
screen "MTA-AyudaVentiladores" 1280x800, template "Plantilla"
   GraphicIOField "Campo ES gráfico_6" at 328,342 size 511x6
   TextField "Campo de texto_5" at 957,566 size 184x61
   TextField "Campo de texto_8" at 218,134 size 461x58
   TextField "Campo de texto_9" at 818,131 size 279x58
   TextField "Campo de texto_1" at 207,101 size 436x42
   TextField "Campo de texto_2" at 807,101 size 179x42
   TextField "Campo de texto_4" at 197,542 size 250x61
   TextField "Campo de texto_7" at 107,251 size 135x42
   GraphicView "Visor de gráficos_3" at 508,439 size 242x85
   GraphicView "Visor de gráficos_4" at 508,253 size 226x85
   GraphicView "Visor de gráficos_5" at 473,452 size 29x29
   GraphicView "Visor de gráficos_6" at 473,268 size 29x29
   TextField "Campo de texto_12" at 957,478 size 156x61
   TextField "Campo de texto_13" at 957,310 size 156x61
   TextField "Campo de texto_3" at 793,372 size 160x42
   TextField "Campo de texto_6" at 413,638 size 729x61
   TextField "Campo de texto_14" at 464,385 size 38x23
   TextField "Campo de texto_15" at 448,209 size 54x23
   TextField "Campo de texto_16" at 556,9 size 171x27
   TextField "Campo de texto_11" at 337,268 size 126x32
   SymbolicIOField "Campo ES simbólico_1" at 339,304 size 170x21
   GraphicIOField "Campo ES gráfico_1" at 328,524 size 511x6
   TextField "Campo de texto_10" at 337,452 size 126x32
   SymbolicIOField "Campo ES simbólico_2" at 339,488 size 170x21
   GraphicView "Visor de gráficos_18" at 757,262 size 71x70
   GraphicView "Visor de gráficos_1" at 757,446 size 71x70
   GraphicView "Visor de gráficos_2" at 757,446 size 71x70

screen "MTA-Booster" 1280x800, template "Plantilla"
   IOField "Campo ES_19" at 28,357 size 90x23
   IOField "Campo ES_17" at 1109,356 size 90x23
   GraphicView "Visor de gráficos_3" at 185,341 size 300x202
   TextField "Campo de texto_16" at 0,10 size 1280x27
   GraphicIOField "Campo ES gráfico_1" at 238,431 size 64x70
   GraphicIOField "Campo ES gráfico_2" at 364,296 size 34x52
   GraphicIOField "Campo ES gráfico_3" at 208,410 size 221x101
   SymbolicIOField "Campo ES simbólico_1" at 949,53 size 322x37
   SymbolicIOField "Campo ES simbólico_2" at 949,95 size 321x37
   GraphicView "Visor de gráficos_4" at 761,341 size 300x202
   GraphicIOField "Campo ES gráfico_4" at 814,431 size 64x70
   GraphicIOField "Campo ES gráfico_5" at 940,296 size 34x52
   GraphicIOField "Campo ES gráfico_6" at 784,410 size 221x101
   GraphicView "Visor de gráficos_2" at 460,408 size 40x40
   GraphicView "Visor de gráficos_1" at 460,408 size 40x40
   Button "Botón_6" at 460,408 size 40x40
   IOField "Campo ES_1" at 217,338 size 90x23
   IOField "Campo ES_2" at 790,338 size 90x23
   Switch "Interruptor_2" at 361,96 size 72x40
   TextField "Campo de texto_1" at 25,103 size 312x23
   Button "Botón_1" at 518,484 size 185x39
   IOField "Campo ES_3" at 359,151 size 130x31
   TextField "Campo de texto_2" at 241,152 size 93x23
   IOField "Campo ES_4" at 359,191 size 130x31
   TextField "Campo de texto_3" at 78,192 size 255x23
   IOField "Campo ES_5" at 359,231 size 130x31
   TextField "Campo de texto_4" at 61,232 size 273x23
   TextField "Campo de texto_5" at 187,550 size 250x27
   TextField "Campo de texto_6" at 762,550 size 250x27
   Button "Botón_7" at 849,639 size 100x27
   Button "Botón_8" at 849,607 size 100x27
   Button "Botón_9" at 960,607 size 96x27
   Button "Botón_10" at 960,639 size 96x27
   Switch "Interruptor_3" at 730,607 size 96x59
   GraphicView "Visor de gráficos_5" at 1036,408 size 40x40
   GraphicView "Visor de gráficos_6" at 1036,408 size 40x40
   Button "Botón_11" at 1036,408 size 40x40
   Button "Botón_2" at 275,639 size 96x27
   Button "Botón_3" at 275,607 size 96x27
   Button "Botón_5" at 384,607 size 96x27
   Button "Botón_4" at 384,639 size 96x27
   Switch "Interruptor_1" at 153,607 size 96x59
   IOField "Campo ES_6" at 217,362 size 90x23
   IOField "Campo ES_7" at 790,362 size 90x23
   IOField "Campo ES_8" at 217,386 size 90x23
   IOField "Campo ES_9" at 790,386 size 90x23
   IOField "Campo ES_10" at 854,140 size 90x23
   IOField "Campo ES_11" at 854,169 size 90x23
   IOField "Campo ES_12" at 854,198 size 90x23
   IOField "Campo ES_13" at 854,227 size 90x23
   IOField "Campo ES_14" at 854,256 size 90x23
   TextField "Campo de texto_7" at 949,140 size 321x139
   TextField "Campo de texto_8" at 187,550 size 250x27
   TextField "Campo de texto_9" at 762,550 size 250x27
   Button "Botón_13" at 985,181 size 96x30
   Button "Botón_14" at 1139,181 size 96x30
   Button "Botón_12" at 985,233 size 252x30
   TrendView "Visor de curvas_1" at 5,53 size 584x236
   TextField "Campo de texto_10" at 591,140 size 241x23
   TextField "Campo de texto_11" at 591,169 size 241x23
   TextField "Campo de texto_12" at 591,198 size 105x23
   TextField "Campo de texto_13" at 591,227 size 259x23
   TextField "Campo de texto_14" at 591,256 size 259x23
   IOField "Campo ES_15" at 854,111 size 90x23
   TextField "Campo de texto_15" at 591,111 size 226x23
   IOField "Campo ES_16" at 854,82 size 90x23
   TextField "Campo de texto_17" at 591,82 size 226x23
   Button "Botón_15" at 49,396 size 96x35
   TextField "Campo de texto_19" at 28,335 size 133x18
   Button "Botón_16" at 1130,395 size 96x35
   TextField "Campo de texto_18" at 1109,334 size 133x18

screen "MTA-CFGALTA" 1280x800, template "Plantilla"
   TextField "Campo de texto_4" at 1016,131 size 91x20
   TextField "Campo de texto_5" at 1016,163 size 84x20
   IOField "Campo ES_4" at 1126,129 size 98x23
   IOField "Campo ES_5" at 1126,161 size 98x23
   TextField "Campo de texto_1" at 49,157 size 275x27
   TextField "Campo de texto_2" at 49,277 size 316x27
   IOField "Campo ES_1" at 630,157 size 130x31
   IOField "Campo ES_2" at 629,277 size 130x31
   TextField "Campo de texto_6" at 49,405 size 526x27
   IOField "Campo ES_3" at 629,405 size 130x31
   TextField "Campo de texto_7" at 902,142 size 94x27
   TextField "Campo de texto_8" at 1016,203 size 91x20
   TextField "Campo de texto_9" at 1016,235 size 84x20
   TextField "Campo de texto_10" at 902,214 size 94x27
   IOField "Campo ES_6" at 1126,201 size 98x23
   IOField "Campo ES_7" at 1126,233 size 98x23
   TextField "Campo de texto_11" at 1016,275 size 91x20
   TextField "Campo de texto_12" at 1016,307 size 84x20
   TextField "Campo de texto_13" at 902,286 size 94x27
   IOField "Campo ES_8" at 1126,273 size 98x23
   IOField "Campo ES_9" at 1126,305 size 98x23
   TextField "Campo de texto_14" at 1016,347 size 91x20
   TextField "Campo de texto_15" at 1016,379 size 84x20
   TextField "Campo de texto_16" at 902,358 size 94x27
   IOField "Campo ES_10" at 1126,345 size 98x23
   IOField "Campo ES_11" at 1126,377 size 98x23
   TextField "Campo de texto_17" at 1016,419 size 91x20
   TextField "Campo de texto_18" at 1016,451 size 84x20
   TextField "Campo de texto_19" at 902,430 size 94x27
   IOField "Campo ES_12" at 1126,417 size 98x23
   IOField "Campo ES_13" at 1126,449 size 98x23
   Button "Botón_12" at 1076,638 size 160x49
   TextField "Campo de texto_3" at 58,190 size 417x22
   TextField "Campo de texto_20" at 58,310 size 566x40
   TextField "Campo de texto_21" at 58,438 size 512x22
   TextField "Campo de texto_22" at 49,509 size 249x27
   TextField "Campo de texto_23" at 58,542 size 542x40
   IOField "Campo ES_14" at 629,509 size 130x31
   TextField "Campo de texto_24" at 1016,563 size 91x20
   TextField "Campo de texto_25" at 1016,595 size 84x20
   TextField "Campo de texto_26" at 902,574 size 55x27
   IOField "Campo ES_15" at 1126,561 size 98x23
   IOField "Campo ES_16" at 1126,593 size 98x23
   Button "Botón_1" at 1184,68 size 48x46
   TextField "Campo de texto_27" at 349,9 size 585x27
   TextField "Campo de texto_28" at 902,502 size 94x27
   TextField "Campo de texto_29" at 1015,491 size 91x20
   TextField "Campo de texto_30" at 1015,523 size 84x20
   IOField "Campo ES_17" at 1125,489 size 98x23
   IOField "Campo ES_18" at 1125,521 size 98x23

screen "MTA-CFGAvisosALTA" 1280x800, template "Plantilla"
   TextField "Campo de texto_1" at 71,96 size 326x27
   TextField "Campo de texto_2" at 683,96 size 276x27
   IOField "Campo ES_1" at 499,96 size 130x31
   IOField "Campo ES_2" at 1110,96 size 130x31
   TextField "Campo de texto_3" at 71,146 size 322x27
   IOField "Campo ES_4" at 498,146 size 130x31
   TextField "Campo de texto_9" at 151,49 size 283x34
   TextField "Campo de texto_4" at 477,9 size 349x27
   TextField "Campo de texto_8" at 71,197 size 397x27
   IOField "Campo ES_5" at 518,197 size 90x23
   TextField "Campo de texto_7" at 683,197 size 397x27
   IOField "Campo ES_6" at 1130,197 size 90x23
   TextField "Campo de texto_10" at 71,246 size 397x27
   IOField "Campo ES_7" at 518,246 size 90x23
   TextField "Campo de texto_11" at 683,246 size 397x27
   IOField "Campo ES_8" at 1130,246 size 90x23
   TextField "Campo de texto_12" at 71,296 size 397x27
   IOField "Campo ES_9" at 518,296 size 90x23
   TextField "Campo de texto_14" at 71,443 size 412x27
   IOField "Campo ES_11" at 518,443 size 90x23
   TextField "Campo de texto_15" at 683,443 size 412x27
   IOField "Campo ES_12" at 1130,443 size 90x23
   TextField "Campo de texto_18" at 683,345 size 397x27
   IOField "Campo ES_15" at 1130,345 size 90x23
   TextField "Campo de texto_19" at 71,393 size 397x27
   IOField "Campo ES_16" at 518,393 size 90x23
   TextField "Campo de texto_20" at 683,296 size 397x27
   IOField "Campo ES_17" at 1130,296 size 90x23
   TextField "Campo de texto_17" at 71,345 size 397x27
   IOField "Campo ES_14" at 518,345 size 90x23
   TextField "Campo de texto_6" at 683,146 size 248x27
   IOField "Campo ES_3" at 1110,146 size 130x31
   TextField "Campo de texto_13" at 683,393 size 397x27
   IOField "Campo ES_10" at 1130,393 size 90x23
   TextField "Campo de texto_5" at 683,590 size 380x27
   Switch "Interruptor_1" at 1155,583 size 37x37
   TextField "Campo de texto_16" at 71,493 size 374x27
   IOField "Campo ES_13" at 518,493 size 90x23
   TextField "Campo de texto_21" at 71,539 size 374x27
   IOField "Campo ES_18" at 518,539 size 90x23
   TextField "Campo de texto_22" at 683,493 size 374x27
   IOField "Campo ES_19" at 1130,493 size 90x23
   TextField "Campo de texto_23" at 683,539 size 390x27
   IOField "Campo ES_20" at 1130,539 size 90x23
   TextField "Campo de texto_31" at 71,589 size 397x27
   IOField "Campo ES_21" at 518,589 size 90x23
   TextField "Campo de texto_24" at 684,637 size 408x27
   Switch "Interruptor_2" at 1156,630 size 37x37

screen "MTA-CFGAvisosBAJA" 1280x800, template "Plantilla"
   TextField "Campo de texto_1" at 477,9 size 354x27
   TextField "Campo de texto_9" at 161,54 size 281x34
   IOField "Campo ES_1" at 295,105 size 130x30
   IOField "Campo ES_2" at 295,240 size 130x31
   IOField "Campo ES_3" at 295,195 size 130x31
   IOField "Campo ES_4" at 295,150 size 130x31
   IOField "Campo ES_5" at 295,285 size 130x30
   IOField "Campo ES_6" at 295,330 size 130x31
   IOField "Campo ES_7" at 295,375 size 130x31
   IOField "Campo ES_8" at 295,420 size 130x31
   TextField "Campo de texto_2" at 15,107 size 293x25
   TextField "Campo de texto_3" at 15,242 size 238x25
   TextField "Campo de texto_6" at 15,197 size 248x25
   TextField "Campo de texto_4" at 15,152 size 289x25
   TextField "Campo de texto_5" at 15,287 size 238x25
   TextField "Campo de texto_7" at 15,332 size 238x25
   TextField "Campo de texto_8" at 15,377 size 238x25
   TextField "Campo de texto_10" at 15,422 size 231x25
   IOField "Campo ES_9" at 295,465 size 130x30
   IOField "Campo ES_10" at 295,510 size 130x31
   IOField "Campo ES_11" at 295,555 size 130x31
   TextField "Campo de texto_11" at 15,467 size 231x25
   TextField "Campo de texto_12" at 15,512 size 231x25
   TextField "Campo de texto_13" at 15,557 size 232x25
   IOField "Campo ES_13" at 716,150 size 130x30
   IOField "Campo ES_14" at 716,105 size 130x31
   IOField "Campo ES_15" at 716,195 size 130x31
   IOField "Campo ES_16" at 716,240 size 130x31
   IOField "Campo ES_17" at 716,285 size 130x30
   IOField "Campo ES_18" at 716,330 size 130x31
   IOField "Campo ES_19" at 716,375 size 130x31
   IOField "Campo ES_20" at 716,420 size 130x31
   TextField "Campo de texto_15" at 436,152 size 248x25
   TextField "Campo de texto_16" at 436,107 size 247x25
   TextField "Campo de texto_17" at 436,197 size 248x25
   TextField "Campo de texto_18" at 436,242 size 238x25
   TextField "Campo de texto_19" at 436,287 size 238x25
   TextField "Campo de texto_20" at 436,332 size 238x25
   TextField "Campo de texto_21" at 436,377 size 231x25
   TextField "Campo de texto_22" at 436,422 size 231x25
   IOField "Campo ES_21" at 716,465 size 130x30
   IOField "Campo ES_22" at 716,510 size 130x31
   IOField "Campo ES_23" at 716,555 size 130x31
   TextField "Campo de texto_23" at 436,467 size 231x25
   TextField "Campo de texto_24" at 436,512 size 231x25
   TextField "Campo de texto_25" at 436,557 size 232x25
   IOField "Campo ES_25" at 1137,195 size 130x30
   IOField "Campo ES_26" at 1137,150 size 130x31
   IOField "Campo ES_27" at 1137,105 size 130x31
   IOField "Campo ES_28" at 1137,240 size 130x31
   IOField "Campo ES_29" at 1137,285 size 130x30
   IOField "Campo ES_30" at 1137,330 size 130x31
   IOField "Campo ES_31" at 1137,375 size 130x31
   IOField "Campo ES_32" at 1137,420 size 130x31
   TextField "Campo de texto_27" at 857,197 size 243x25
   TextField "Campo de texto_28" at 857,152 size 248x25
   TextField "Campo de texto_29" at 857,107 size 222x25
   TextField "Campo de texto_30" at 857,242 size 238x25
   TextField "Campo de texto_31" at 857,287 size 238x25
   TextField "Campo de texto_32" at 857,332 size 238x25
   TextField "Campo de texto_33" at 857,377 size 231x25
   TextField "Campo de texto_34" at 857,422 size 273x25
   IOField "Campo ES_33" at 1137,465 size 130x30
   IOField "Campo ES_34" at 1137,510 size 130x31
   IOField "Campo ES_35" at 1137,555 size 130x31
   TextField "Campo de texto_35" at 857,467 size 231x25
   TextField "Campo de texto_36" at 857,512 size 232x25
   TextField "Campo de texto_37" at 857,557 size 232x25

screen "MTA-ChillersBombasEnvasado" 1280x800, template "Plantilla"
   TextField "Campo de texto_5" at 519,10 size 240x27
   GraphicView "Visor de gráficos_3" at 944,375 size 64x103
   GraphicIOField "Plantilla_Campo ES gráfico_2" at 980,449 size 81x68
   SymbolicIOField "Campo ES simbólico_4" at 890,188 size 220x29
   TextField "Campo de texto_6" at 887,129 size 53x23
   GraphicView "Visor de gráficos_4" at 702,375 size 64x103
   GraphicIOField "Plantilla_Campo ES gráfico_1" at 738,449 size 81x68
   SymbolicIOField "Campo ES simbólico_1" at 648,188 size 220x29
   TextField "Campo de texto_7" at 645,129 size 53x23
   GraphicView "Visor de gráficos_6" at 216,375 size 64x103
   GraphicIOField "Plantilla_Campo ES gráfico_4" at 252,449 size 81x68
   SymbolicIOField "Campo ES simbólico_3" at 164,188 size 220x29
   TextField "Campo de texto_9" at 167,129 size 52x23
   TextField "Campo de texto_19" at 645,160 size 195x18
   GraphicView "Visor de gráficos_5" at 460,375 size 64x103
   GraphicIOField "Plantilla_Campo ES gráfico_3" at 496,449 size 81x68
   SymbolicIOField "Campo ES simbólico_2" at 406,188 size 220x29
   TextField "Campo de texto_8" at 403,129 size 52x23
   TextField "Campo de texto_18" at 886,160 size 150x18
   TextField "Campo de texto_16" at 407,161 size 150x18
   TextField "Campo de texto_17" at 165,161 size 146x18
   ScreenModuleView "ControlMotor-NoAUTO_1" at 916,230 size 171x108
   ScreenModuleView "ControlMotor-NoAUTO_2" at 676,230 size 171x108
   ScreenModuleView "ControlMotor-NoAUTO_3" at 431,230 size 171x108
   ScreenModuleView "ControlMotor-NoAUTO_4" at 191,230 size 171x108
   Button "Botón_1" at 1184,68 size 48x46

screen "MTA-ChillersBombasSoplado" 1280x800, template "Plantilla"
   GraphicView "Visor de gráficos_3" at 944,375 size 64x103
   GraphicView "Visor de gráficos_4" at 702,375 size 64x103
   GraphicView "Visor de gráficos_6" at 216,375 size 64x103
   GraphicView "Visor de gráficos_5" at 460,375 size 64x103
   TextField "Campo de texto_5" at 530,10 size 221x27
   GraphicIOField "Plantilla_Campo ES gráfico_2" at 980,449 size 81x68
   SymbolicIOField "Campo ES simbólico_4" at 890,188 size 220x29
   TextField "Campo de texto_6" at 887,129 size 53x23
   GraphicIOField "Plantilla_Campo ES gráfico_1" at 738,449 size 81x68
   SymbolicIOField "Campo ES simbólico_1" at 648,188 size 220x29
   TextField "Campo de texto_7" at 645,129 size 53x23
   GraphicIOField "Plantilla_Campo ES gráfico_4" at 252,449 size 81x68
   SymbolicIOField "Campo ES simbólico_3" at 164,188 size 220x29
   TextField "Campo de texto_9" at 167,129 size 52x23
   TextField "Campo de texto_19" at 647,161 size 166x18
   GraphicIOField "Plantilla_Campo ES gráfico_3" at 496,449 size 81x68
   SymbolicIOField "Campo ES simbólico_2" at 406,188 size 220x29
   TextField "Campo de texto_8" at 403,129 size 52x23
   TextField "Campo de texto_18" at 887,161 size 104x18
   TextField "Campo de texto_16" at 404,161 size 142x18
   TextField "Campo de texto_17" at 165,161 size 138x18
   GraphicView "Plantilla_Visor de gráficos_2" at 1232,6 size 35x35
   GraphicView "Plantilla_Visor de gráficos_1" at 1232,6 size 35x35
   Button "Botón_1" at 1220,1 size 57x44
   ScreenModuleView "ControlMotor-NoAUTO_4" at 916,230 size 171x108
   ScreenModuleView "ControlMotor-NoAUTO_1" at 424,229 size 171x108
   ScreenModuleView "ControlMotor-NoAUTO_2" at 676,230 size 171x108
   ScreenModuleView "ControlMotor-NoAUTO_3" at 184,229 size 171x108
   Button "Botón_2" at 1184,68 size 48x46

screen "MTA-ChillersCFGSirena" 1280x800, template "Plantilla"
   Switch "Interruptor_1" at 215,155 size 36x32
   Switch "Interruptor_2" at 215,192 size 36x32
   Switch "Interruptor_3" at 215,229 size 36x32
   Switch "Interruptor_4" at 215,266 size 36x32
   Switch "Interruptor_5" at 215,303 size 36x32
   TextField "Campo de texto_1" at 259,307 size 365x22
   TextField "Campo de texto_2" at 259,270 size 424x22
   TextField "Campo de texto_3" at 259,234 size 353x22
   TextField "Campo de texto_4" at 259,196 size 411x22
   TextField "Campo de texto_5" at 259,160 size 340x22
   TextField "Campo de texto_6" at 147,93 size 410x22
   Switch "Interruptor_6" at 215,340 size 36x32
   TextField "Campo de texto_8" at 259,345 size 231x22
   Switch "Interruptor_7" at 215,377 size 36x32
   TextField "Campo de texto_9" at 259,381 size 244x22
   Switch "Interruptor_8" at 215,415 size 36x32
   TextField "Campo de texto_10" at 259,420 size 150x22
   GraphicView "Plantilla_Visor de gráficos_2" at 1232,6 size 35x35
   GraphicView "Plantilla_Visor de gráficos_1" at 1232,6 size 35x35
   Button "Botón_1" at 1220,1 size 57x44
   Switch "Interruptor_9" at 215,453 size 36x32
   TextField "Campo de texto_11" at 259,458 size 194x22
   TextField "Campo de texto_7" at 505,9 size 270x27

screen "MTA-Chillers-General" 1280x800, template "Plantilla"
   GraphicView "Visor de gráficos_7" at 774,285 size 48x87
   GraphicView "Visor de gráficos_8" at 838,285 size 48x87
   GraphicView "Visor de gráficos_1" at 646,285 size 48x87
   GraphicView "Visor de gráficos_9" at 710,285 size 48x87
   GraphicView "Visor de gráficos_3" at 1155,429 size 120x284
   GraphicView "Visor de gráficos_4" at 950,233 size 168x168
   GraphicView "Visor de gráficos_5" at 494,285 size 48x87
   GraphicView "Visor de gráficos_6" at 558,285 size 48x87
   GraphicView "Visor de gráficos_10" at 366,285 size 48x87
   GraphicView "Visor de gráficos_11" at 430,285 size 48x87
   GraphicView "Visor de gráficos_2" at 12,188 size 200x216
   GraphicView "Visor de gráficos_12" at 107,550 size 160x149
   GraphicView "Visor de gráficos_15" at 351,213 size 116x103
   GraphicView "Visor de gráficos_16" at 479,213 size 116x103
   GraphicView "Visor de gráficos_17" at 631,213 size 116x103
   GraphicView "Visor de gráficos_18" at 759,213 size 116x103
   GraphicView "Visor de gráficos_14" at 622,54 size 245x227
   GraphicView "Visor de gráficos_13" at 344,46 size 245x227
   GraphicView "Plantilla_Visor de gráficos_2" at 1232,6 size 35x35
   GraphicView "Plantilla_Visor de gráficos_1" at 1232,6 size 35x35
   GraphicIOField "Plantilla_Campo ES gráfico_2" at 529,355 size 57x52
   GraphicIOField "Plantilla_Campo ES gráfico_1" at 593,355 size 57x52
   GraphicIOField "Plantilla_Campo ES gráfico_3" at 809,355 size 57x52
   GraphicIOField "Plantilla_Campo ES gráfico_4" at 873,355 size 57x52
   GraphicIOField "Plantilla_Campo ES gráfico_5" at 681,355 size 57x52
   GraphicIOField "Plantilla_Campo ES gráfico_6" at 745,355 size 57x52
   GraphicIOField "Plantilla_Campo ES gráfico_7" at 401,355 size 57x52
   GraphicIOField "Plantilla_Campo ES gráfico_8" at 465,355 size 57x52
   TextField "Campo de texto_1" at 984,196 size 86x32
   TextField "Campo de texto_2" at 1027,485 size 86x32
   TextField "Campo de texto_3" at 134,514 size 90x32
   TextField "Campo de texto_4" at 60,150 size 90x32
   TextField "Campo de texto_6" at 762,451 size 131x25
   TextField "Campo de texto_7" at 477,451 size 139x25
   TextField "Campo de texto_9" at 848,132 size 51x52
   TextField "Campo de texto_8" at 424,419 size 41x19
   TextField "Campo de texto_11" at 485,419 size 41x19
   TextField "Campo de texto_12" at 546,419 size 49x19
   TextField "Campo de texto_13" at 614,419 size 42x19
   TextField "Campo de texto_14" at 703,419 size 41x19
   TextField "Campo de texto_15" at 767,419 size 41x19
   TextField "Campo de texto_16" at 830,419 size 42x19
   TextField "Campo de texto_17" at 893,419 size 42x19
   TextField "Campo de texto_10" at 569,131 size 58x52
   TextField "Campo de texto_21" at 242,362 size 40x18
   TextField "Campo de texto_22" at 242,341 size 108x18
   TextField "Campo de texto_23" at 242,382 size 101x18
   TextField "Campo de texto_24" at 299,638 size 79x18
   TextField "Campo de texto_25" at 299,617 size 108x18
   TextField "Campo de texto_26" at 299,660 size 115x18
   TextField "Campo de texto_27" at 299,681 size 125x18
   TextField "Campo de texto_18" at 1037,602 size 40x18
   TextField "Campo de texto_19" at 1037,581 size 108x18
   TextField "Campo de texto_20" at 1037,622 size 101x18
   TextField "Campo de texto_28" at 1154,313 size 120x18
   TextField "Campo de texto_29" at 1154,292 size 120x18
   TextField "Campo de texto_30" at 1154,335 size 96x18
   TextField "Campo de texto_31" at 1154,356 size 96x18
   Button "Botón_2" at 657,329 size 295x86
   Button "Botón_5" at 361,328 size 296x87
   Button "Botón_1" at 1220,1 size 57x44
   Switch "Interruptor_1" at 222,294 size 91x31
   Switch "Interruptor_2" at 279,570 size 91x31
   Switch "Interruptor_3" at 1017,534 size 91x31
   Switch "Interruptor_4" at 1135,252 size 91x31
   Button "Botón_3" at 1184,68 size 48x46
   TextField "Campo de texto_32" at 610,9 size 63x27

screen "MTA-CompBAJA" 1280x800, template "Plantilla"
   GraphicIOField "Campo ES gráfico_10" at 360,303 size 189x58
   GraphicIOField "Campo ES gráfico_9" at 296,391 size 189x58
   GraphicIOField "Campo ES gráfico_8" at 524,183 size 197x58
   GraphicView "Visor de gráficos_1" at 336,222 size 269x127
   GraphicView "Visor de gráficos_7" at 336,222 size 269x127
   GraphicView "Visor de gráficos_2" at 272,310 size 269x127
   GraphicView "Visor de gráficos_8" at 272,310 size 269x127
   GraphicView "Visor de gráficos_5" at 506,105 size 213x127
   GraphicView "Visor de gráficos_11" at 506,105 size 213x127
   GraphicView "Visor de gráficos_6" at 132,415 size 202x177
   IOField "Campo ES_1" at 160,512 size 148x28
   Button "Botón_3" at 1184,48 size 48x46
   Button "Botón_1" at 35,197 size 160x46
   TextField "Campo de texto_1" at 516,9 size 248x27
   GraphicIOField "Campo ES gráfico_1" at 581,409 size 507x6
   GraphicIOField "Campo ES gráfico_4" at 769,184 size 511x6
   GraphicIOField "Campo ES gráfico_5" at 630,322 size 507x6
   TextField "Campo de texto_5" at 794,109 size 116x39
   TextField "Campo de texto_8" at 598,335 size 91x39
   TextField "Campo de texto_9" at 654,247 size 100x39
   SymbolicIOField "Campo ES simbólico_5" at 656,283 size 242x21
   SymbolicIOField "Campo ES simbólico_6" at 600,371 size 242x21
   SymbolicIOField "Campo ES simbólico_9" at 796,145 size 242x21
   IOField "Campo ES_6" at 796,165 size 85x19
   IOField "Campo ES_7" at 600,390 size 85x19
   IOField "Campo ES_8" at 656,302 size 85x19
   Switch "Interruptor_1" at 852,252 size 29x29
   Switch "Interruptor_2" at 802,340 size 29x29
   ScreenModuleView "Faceplate_1_4" at 849,342 size 236x58
   ScreenModuleView "Faceplate_1_5" at 899,255 size 236x58
   Switch "Interruptor_7" at 402,135 size 40x40
   Switch "Interruptor_9" at 234,321 size 40x40
   Switch "Interruptor_10" at 298,233 size 40x40
   Switch "Interruptor_5" at 1131,132 size 91x31
   Button "Botón_14" at 769,109 size 262x74
   Button "Botón_17" at 581,335 size 200x74
   Button "Botón_18" at 629,247 size 200x74

screen "MTA-SecALTA" 1280x800, template "Plantilla"
   GraphicIOField "Campo ES gráfico_4" at 981,258 size 280x222
   GraphicView "Visor de gráficos_4" at 999,137 size 234x314
   GraphicView "Visor de gráficos_15" at 999,137 size 234x314
   GraphicIOField "Campo ES gráfico_8" at 571,212 size 366x99
   GraphicView "Visor de gráficos_3" at 592,100 size 363x184
   GraphicView "Visor de gráficos_5" at 592,100 size 363x184
   GraphicIOField "Campo ES gráfico_7" at 674,357 size 309x81
   GraphicView "Visor de gráficos_2" at 696,255 size 292x158
   GraphicView "Visor de gráficos_6" at 695,255 size 294x158
   GraphicIOField "Campo ES gráfico_6" at 765,490 size 338x86
   GraphicView "Visor de gráficos_1" at 786,405 size 292x142
   GraphicView "Visor de gráficos_14" at 786,405 size 292x142
   Button "Botón_3" at 1184,68 size 48x46
   TextField "Campo de texto_7" at 530,9 size 221x27
   GraphicIOField "Campo ES gráfico_9" at 197,577 size 511x6
   TextField "Campo de texto_6" at 222,499 size 89x39
   SymbolicIOField "Campo ES simbólico_9" at 224,535 size 242x21
   GraphicIOField "Campo ES gráfico_1" at 101,439 size 511x6
   TextField "Campo de texto_1" at 126,361 size 89x39
   SymbolicIOField "Campo ES simbólico_1" at 128,397 size 242x21
   GraphicIOField "Campo ES gráfico_2" at 21,303 size 511x6
   TextField "Campo de texto_2" at 46,220 size 101x39
   SymbolicIOField "Campo ES simbólico_2" at 48,256 size 242x21
   GraphicIOField "Campo ES gráfico_3" at 741,681 size 511x6
   TextField "Campo de texto_3" at 766,603 size 89x39
   SymbolicIOField "Campo ES simbólico_3" at 768,639 size 242x21
   IOField "Campo ES_6" at 51,282 size 85x19
   IOField "Campo ES_1" at 131,418 size 85x19
   IOField "Campo ES_2" at 227,558 size 85x19
   IOField "Campo ES_3" at 771,660 size 85x19
   Switch "Interruptor_1" at 640,315 size 40x40
   Switch "Interruptor_2" at 731,440 size 40x40
   Switch "Interruptor_3" at 540,176 size 40x40
   Switch "Interruptor_4" at 1212,488 size 40x40
   Switch "Interruptor_5" at 387,506 size 29x29
   Switch "Interruptor_6" at 307,370 size 29x29
   Switch "Interruptor_7" at 227,229 size 29x29
   Switch "Interruptor_8" at 925,606 size 29x29
   ScreenModuleView "Faceplate_2_1" at 453,489 size 244x69
   ScreenModuleView "Faceplate_2_2" at 357,351 size 244x69
   ScreenModuleView "Faceplate_2_3" at 276,215 size 244x69
   ScreenModuleView "Faceplate_2_4" at 994,593 size 244x69
   Button "Botón_1" at 741,590 size 150x90
   Button "Botón_2" at 197,486 size 150x90
   Button "Botón_4" at 101,348 size 150x90
   Button "Botón_5" at 21,212 size 150x90

screen "MTA-SecBaja" 1280x800, template "Plantilla"
   GraphicIOField "Campo ES gráfico_4" at 639,360 size 511x6
   TextField "Campo de texto_5" at 664,282 size 116x39
   SymbolicIOField "Campo ES simbólico_9" at 666,318 size 242x21
   GraphicIOField "Campo ES gráfico_3" at 482,493 size 510x6
   TextField "Campo de texto_6" at 507,415 size 116x39
   SymbolicIOField "Campo ES simbólico_8" at 509,451 size 242x21
   IOField "Campo ES_6" at 666,339 size 85x19
   IOField "Campo ES_1" at 509,472 size 85x19
   ScreenModuleView "Faceplate_3_2" at 923,282 size 213x73
   ScreenModuleView "Faceplate_3_1" at 761,415 size 213x73
   Switch "Interruptor_7" at 271,262 size 40x40
   Switch "Interruptor_8" at 131,406 size 40x40
   GraphicIOField "Campo ES gráfico_1" at 289,314 size 285x90
   GraphicView "Visor de gráficos_2" at 333,200 size 201x179
   GraphicIOField "Campo ES gráfico_8" at 159,455 size 269x90
   GraphicView "Visor de gráficos_4" at 333,200 size 201x179
   GraphicView "Visor de gráficos_1" at 192,341 size 201x179
   GraphicView "Visor de gráficos_3" at 192,341 size 201x179
   Button "Botón_3" at 1184,68 size 48x46
   TextField "Campo de texto_1" at 527,9 size 226x27
   Button "Botón_18" at 639,277 size 200x82
   Button "Botón_1" at 482,410 size 200x82

screen "MTA-Sopladoras" 1280x800, template "Plantilla"
   IOField "Campo ES_1" at 301,378 size 151x31
   IOField "Campo ES_2" at 492,378 size 153x31
   IOField "Campo ES_3" at 691,378 size 153x31
   IOField "Campo ES_4" at 766,443 size 90x23
   TextField "Campo de texto_1" at 356,442 size 403x27
   TextField "Campo de texto_2" at 328,211 size 104x27
   Button "Botón_12" at 1105,638 size 160x49
   Button "Botón_1" at 323,269 size 112x38
   Button "Botón_2" at 323,309 size 112x38
   Button "Botón_3" at 513,269 size 112x38
   Button "Botón_4" at 513,309 size 112x38
   Button "Botón_5" at 711,269 size 112x38
   Button "Botón_6" at 711,309 size 112x38
   TextField "Campo de texto_3" at 518,211 size 104x27
   TextField "Campo de texto_4" at 716,211 size 104x27
   TextField "Campo de texto_7" at 522,9 size 236x27

screen "MTA-TiemposCmpAlta" 1280x800, template "Plantilla"
   TextField "Campo de texto_3" at 278,160 size 235x27
   IOField "Campo ES_5" at 889,160 size 90x23
   TextField "Campo de texto_1" at 278,288 size 268x27
   IOField "Campo ES_1" at 889,288 size 90x23
   TextField "Campo de texto_2" at 278,432 size 339x27
   IOField "Campo ES_2" at 889,432 size 90x23
   TextField "Campo de texto_4" at 286,192 size 586x36
   TextField "Campo de texto_5" at 286,320 size 616x52
   TextField "Campo de texto_6" at 286,464 size 578x36
   Button "Botón_12" at 1105,638 size 160x49
   TextField "Campo de texto_7" at 477,9 size 326x27

screen "MTA-TorresCAV" 1280x800, template "Plantilla"
   GraphicView "Visor de gráficos_9" at 71,137 size 234x255
   GraphicView "Visor de gráficos_11" at 71,137 size 234x255
   GraphicView "Visor de gráficos_14" at 71,137 size 234x255
   GraphicView "Visor de gráficos_1" at 271,121 size 282x311
   GraphicView "Visor de gráficos_2" at 271,121 size 282x311
   GraphicView "Visor de gráficos_3" at 271,121 size 282x311
   ScreenModuleView "Faceplate_9_2" at 831,282 size 221x68
   ScreenModuleView "Faceplate_9_1" at 831,173 size 221x68
   GraphicView "Visor de gráficos_17" at 7,412 size 77x78
   GraphicView "Visor de gráficos_16" at 340,421 size 190x41
   TextField "Campo de texto_23" at 647,286 size 126x32
   TextField "Campo de texto_3" at 647,178 size 126x32
   GraphicIOField "Campo ES gráfico_4" at 638,358 size 511x6
   GraphicIOField "Campo ES gráfico_5" at 638,250 size 511x6
   SymbolicIOField "Campo ES simbólico_6" at 649,322 size 170x21
   SymbolicIOField "Campo ES simbólico_2" at 649,214 size 170x21
   Switch "Interruptor_5" at 782,288 size 29x29
   Switch "Interruptor_1" at 782,180 size 29x29
   GraphicIOField "Campo ES gráfico_8" at 798,700 size 418x6
   GraphicIOField "Campo ES gráfico_9" at 52,700 size 418x6
   TextField "Campo de texto_8" at 815,623 size 155x32
   TextField "Campo de texto_9" at 64,623 size 182x32
   SymbolicIOField "Campo ES simbólico_5" at 817,659 size 170x21
   SymbolicIOField "Campo ES simbólico_7" at 73,659 size 170x21
   GraphicView "Visor de gráficos_22" at 1067,281 size 71x70
   GraphicView "Visor de gráficos_23" at 1067,281 size 71x70
   GraphicView "Visor de gráficos_20" at 1067,173 size 71x70
   GraphicView "Visor de gráficos_21" at 1067,173 size 71x70
   ScreenModuleView "ControlMotor-NoAUTO_4" at 1005,625 size 203x65
   ScreenModuleView "ControlMotor-NoAUTO_5" at 259,625 size 203x65
   GraphicView "Visor de gráficos_10" at 511,450 size 13x105
   GraphicView "Visor de gráficos_12" at 625,530 size 14x25
   TextField "Campo de texto_2" at 124,104 size 101x20
   TextField "Campo de texto_1" at 357,88 size 104x23
   GraphicView "Visor de gráficos_13" at 514,528 size 125x10
   GraphicView "Visor de gráficos_7" at 497,527 size 72x111
   GraphicView "Visor de gráficos_8" at 612,527 size 72x111
   TextField "Campo de texto_7" at 697,691 size 48x22
   TextField "Campo de texto_6" at 582,691 size 48x22
   TextField "Campo de texto_4" at 113,471 size 84x27
   GraphicIOField "Plantilla_Campo ES gráfico_2" at 663,615 size 81x68
   GraphicIOField "Plantilla_Campo ES gráfico_1" at 546,615 size 81x68
   TextField "Campo de texto_22" at 661,479 size 90x22
   IOField "Campo ES_7" at 657,499 size 98x23
   GraphicView "Visor de gráficos_33" at 201,338 size 118x71
   GraphicView "Visor de gráficos_4" at 188,396 size 185x41
   GraphicView "Visor de gráficos_5" at 108,374 size 169x37
   GraphicView "Visor de gráficos_6" at 174,385 size 169x37
   GraphicView "Visor de gráficos_15" at 62,386 size 130x79
   Button "Botón_3" at 1184,68 size 48x46
   TextField "Campo de texto_10" at 505,10 size 271x27
   GraphicIOField "Campo ES gráfico_2" at 149,135 size 76x32
   GraphicIOField "Campo ES gráfico_1" at 366,121 size 87x34

screen "MTA-TorresCH" 1280x800, template "Plantilla"
   TextField "Campo de texto_13" at 60,454 size 73x22
   TextField "Campo de texto_7" at 697,691 size 48x22
   TextField "Campo de texto_6" at 582,691 size 48x22
   GraphicView "Visor de gráficos_7" at 497,527 size 72x111
   GraphicView "Plantilla_Visor de gráficos_2" at 1232,6 size 35x35
   GraphicView "Plantilla_Visor de gráficos_1" at 1232,6 size 35x35
   GraphicView "Visor de gráficos_8" at 612,527 size 72x111
   Button "Botón_1" at 1220,1 size 57x44
   GraphicIOField "Plantilla_Campo ES gráfico_2" at 663,615 size 81x68
   GraphicIOField "Plantilla_Campo ES gráfico_1" at 546,615 size 81x68
   TextField "Campo de texto_22" at 661,479 size 90x22
   Button "Botón_3" at 1184,68 size 48x46
   GraphicView "Visor de gráficos_9" at 96,443 size 233x53
   GraphicView "Visor de gráficos_11" at 62,461 size 154x79
   GraphicView "Visor de gráficos_25" at 305,367 size 233x53
   GraphicView "Visor de gráficos_26" at 313,379 size 233x53
   GraphicView "Visor de gráficos_28" at 413,396 size 233x53
   TextField "Campo de texto_10" at 511,10 size 260x27
   IOField "Campo ES_1" at 668,499 size 80x23
   GraphicView "Visor de gráficos_1" at 271,137 size 234x255
   GraphicView "Visor de gráficos_17" at 34,97 size 370x377
   GraphicView "Visor de gráficos_2" at 271,137 size 234x255
   GraphicView "Visor de gráficos_5" at 34,97 size 370x377
   GraphicView "Visor de gráficos_6" at 271,137 size 234x255
   GraphicView "Visor de gráficos_16" at 34,97 size 370x377
   TextField "Campo de texto_2" at 364,104 size 47x20
   TextField "Campo de texto_12" at 188,63 size 57x23
   GraphicView "Visor de gráficos_10" at 511,530 size 13x27
   GraphicView "Visor de gráficos_12" at 625,437 size 14x117
   GraphicView "Visor de gráficos_13" at 511,523 size 118x10
   TextField "Campo de texto_1" at 589,92 size 57x23
   GraphicView "Visor de gráficos_4" at 476,127 size 290x297
   GraphicView "Visor de gráficos_3" at 476,127 size 290x297
   GraphicView "Visor de gráficos_15" at 476,127 size 290x297
   ScreenModuleView "ControlMotor-NoAUTO_4" at 1021,625 size 203x65
   ScreenModuleView "ControlMotor-NoAUTO_5" at 243,625 size 203x65
   GraphicIOField "Campo ES gráfico_1" at 157,95 size 116x44
   GraphicIOField "Campo ES gráfico_2" at 349,135 size 76x32
   GraphicIOField "Campo ES gráfico_3" at 573,122 size 91x39
   GraphicIOField "Campo ES gráfico_4" at 758,214 size 511x6
   TextField "Campo de texto_23" at 767,142 size 126x32
   SymbolicIOField "Campo ES simbólico_6" at 769,178 size 170x21
   Switch "Interruptor_5" at 902,144 size 29x29
   GraphicIOField "Campo ES gráfico_5" at 758,326 size 511x6
   TextField "Campo de texto_3" at 767,254 size 126x32
   SymbolicIOField "Campo ES simbólico_2" at 769,290 size 170x21
   Switch "Interruptor_1" at 902,256 size 29x29
   GraphicIOField "Campo ES gráfico_6" at 758,438 size 511x6
   TextField "Campo de texto_4" at 767,366 size 126x32
   SymbolicIOField "Campo ES simbólico_3" at 769,402 size 170x21
   Switch "Interruptor_2" at 902,368 size 29x29
   TextField "Campo de texto_8" at 831,623 size 155x32
   SymbolicIOField "Campo ES simbólico_5" at 833,659 size 170x21
   TextField "Campo de texto_9" at 47,623 size 182x32
   SymbolicIOField "Campo ES simbólico_7" at 57,659 size 170x21
   GraphicIOField "Campo ES gráfico_8" at 814,700 size 418x6
   GraphicIOField "Campo ES gráfico_9" at 36,700 size 418x6
   ScreenModuleView "Faceplate_9_1" at 950,138 size 221x68
   ScreenModuleView "Faceplate_9_2" at 950,250 size 221x68
   ScreenModuleView "Faceplate_9_3" at 950,362 size 221x68
   GraphicView "Visor de gráficos_22" at 1187,137 size 71x70
   GraphicView "Visor de gráficos_23" at 1187,137 size 71x70
   GraphicView "Visor de gráficos_18" at 1187,360 size 71x70
   GraphicView "Visor de gráficos_19" at 1187,360 size 71x70
   GraphicView "Visor de gráficos_20" at 1187,249 size 71x70
   GraphicView "Visor de gráficos_21" at 1187,249 size 71x70
   GraphicView "Visor de gráficos_14" at 1,492 size 85x70
   GraphicView "Visor de gráficos_24" at 309,399 size 237x95

screen "SentronPAC-MTA" 1280x800, template "Plantilla"
   TextField "Campo de texto_5" at 551,10 size 179x27
   TextField "Campo de texto_4" at 105,133 size 55x27
   TextField "Campo de texto_6" at 337,133 size 54x27
   TextField "Campo de texto_7" at 209,133 size 68x27
   TextField "Campo de texto_14" at 41,165 size 16x27
   IOField "Campo ES_1" at 74,165 size 110x27
   IOField "Campo ES_2" at 74,197 size 110x27
   IOField "Campo ES_3" at 74,229 size 110x27
   IOField "Campo ES_4" at 314,165 size 110x27
   IOField "Campo ES_5" at 194,165 size 110x27
   IOField "Campo ES_6" at 194,197 size 110x27
   IOField "Campo ES_7" at 194,229 size 110x27
   IOField "Campo ES_8" at 74,286 size 110x27
   IOField "Campo ES_9" at 74,318 size 110x27
   IOField "Campo ES_10" at 74,350 size 110x27
   IOField "Campo ES_11" at 314,286 size 110x27
   IOField "Campo ES_12" at 194,286 size 110x27
   IOField "Campo ES_13" at 194,318 size 110x27
   IOField "Campo ES_14" at 194,350 size 110x27
   TextField "Campo de texto_15" at 41,197 size 15x27
   TextField "Campo de texto_16" at 41,229 size 15x27
   TextField "Campo de texto_17" at 41,286 size 27x27
   TextField "Campo de texto_18" at 41,318 size 26x27
   TextField "Campo de texto_19" at 41,350 size 27x27
   TextField "Campo de texto_8" at 105,453 size 55x27
   TextField "Campo de texto_9" at 337,453 size 54x27
   TextField "Campo de texto_10" at 209,453 size 68x27
   TextField "Campo de texto_11" at 41,485 size 16x27
   TextField "Campo de texto_12" at 41,517 size 15x27
   TextField "Campo de texto_13" at 41,549 size 15x27
   IOField "Campo ES_15" at 74,485 size 110x27
   IOField "Campo ES_16" at 74,517 size 110x27
   IOField "Campo ES_17" at 74,549 size 110x27
   IOField "Campo ES_18" at 314,485 size 110x27
   IOField "Campo ES_19" at 194,485 size 110x27
   IOField "Campo ES_20" at 194,517 size 110x27
   IOField "Campo ES_23" at 194,549 size 110x27
   TextField "Campo de texto_20" at 719,133 size 64x27
   TextField "Campo de texto_21" at 703,165 size 16x27
   IOField "Campo ES_24" at 725,165 size 62x27
   TextField "Campo de texto_22" at 703,197 size 15x27
   IOField "Campo ES_25" at 725,197 size 62x27
   TextField "Campo de texto_23" at 703,229 size 15x27
   IOField "Campo ES_26" at 725,229 size 62x27
   TextField "Campo de texto_24" at 671,293 size 45x27
   IOField "Campo ES_27" at 725,293 size 62x27
   TextField "Campo de texto_25" at 823,133 size 53x27
   TextField "Campo de texto_26" at 942,133 size 74x27
   IOField "Campo ES_28" at 797,165 size 126x27
   IOField "Campo ES_29" at 797,197 size 126x27
   IOField "Campo ES_30" at 797,229 size 126x27
   IOField "Campo ES_31" at 931,165 size 126x27
   IOField "Campo ES_32" at 931,197 size 126x27
   IOField "Campo ES_33" at 931,229 size 126x27
   TextField "Campo de texto_27" at 1077,133 size 80x27
   IOField "Campo ES_34" at 1067,165 size 121x27
   IOField "Campo ES_35" at 1067,197 size 121x27
   IOField "Campo ES_36" at 1067,229 size 121x27
   IOField "Campo ES_21" at 797,293 size 126x27
   IOField "Campo ES_22" at 931,293 size 126x27
   IOField "Campo ES_37" at 1067,293 size 121x27
   TextField "Campo de texto_30" at 695,461 size 95x27
   TextField "Campo de texto_31" at 695,493 size 171x27
   TextField "Campo de texto_32" at 695,525 size 182x27
   IOField "Campo ES_38" at 893,461 size 110x27
   IOField "Campo ES_39" at 893,493 size 110x27
   IOField "Campo ES_40" at 893,525 size 110x27
   TextField "Campo de texto_29" at 465,133 size 41x27
   TextField "Campo de texto_33" at 465,453 size 41x27
   IOField "Campo ES_41" at 434,165 size 110x27
   IOField "Campo ES_42" at 434,197 size 110x27
   IOField "Campo ES_43" at 434,229 size 110x27
   IOField "Campo ES_47" at 434,485 size 110x27
   IOField "Campo ES_48" at 434,517 size 110x27
   IOField "Campo ES_49" at 434,549 size 110x27
   TextField "Campo de texto_34" at 31,100 size 603x27
   TextField "Campo de texto_35" at 31,420 size 603x27
   TextField "Campo de texto_1" at 650,100 size 609x27
   TextField "Campo de texto_2" at 655,420 size 601x27
   Button "Botón_1" at 565,186 size 50x49
   Button "Botón_2" at 565,315 size 50x49
   Button "Botón_3" at 565,506 size 50x49
   Button "Botón_4" at 1197,186 size 50x49
   Button "Botón_5" at 1197,282 size 50x49

screen "MTA-AyudaCmpBaja" 1280x800, template "Plantilla"
   GraphicIOField "Campo ES gráfico_7" at 279,380 size 178x52
   GraphicIOField "Campo ES gráfico_1" at 351,380 size 178x52
   GraphicView "Visor de gráficos_3" at 269,294 size 269x127
   GraphicView "Visor de gráficos_9" at 335,168 size 269x127
   TextField "Campo de texto_11" at 50,259 size 199x76
   TextField "Campo de texto_12" at 39,229 size 210x42
   TextField "Campo de texto_2" at 145,116 size 210x42
   TextField "Campo de texto_8" at 762,110 size 352x94
   TextField "Campo de texto_9" at 946,227 size 230x76
   TextField "Campo de texto_4" at 751,85 size 203x42
   TextField "Campo de texto_13" at 991,455 size 195x42
   GraphicView "Visor de gráficos_5" at 920,329 size 202x77
   GraphicIOField "Campo ES gráfico_2" at 621,403 size 507x6
   TextField "Campo de texto_14" at 589,454 size 160x42
   TextField "Campo de texto_15" at 615,261 size 108x61
   GraphicView "Visor de gráficos_1" at 804,336 size 31x31
   TextField "Campo de texto_1" at 789,269 size 54x42
   TextField "Campo de texto_16" at 335,457 size 134x42
   GraphicView "Visor de gráficos_4" at 920,497 size 202x77
   GraphicIOField "Campo ES gráfico_3" at 621,571 size 507x6
   GraphicView "Visor de gráficos_2" at 806,505 size 31x31
   TextField "Campo de texto_17" at 798,443 size 38x42
   TextField "Campo de texto_6" at 477,590 size 726x99
   TextField "Campo de texto_5" at 29,520 size 471x213
   TextField "Campo de texto_10" at 529,9 size 246x27
   TextField "Campo de texto_7" at 645,334 size 116x39
   SymbolicIOField "Campo ES simbólico_7" at 647,370 size 242x21
   TextField "Campo de texto_3" at 645,502 size 116x39
   SymbolicIOField "Campo ES simbólico_1" at 647,538 size 242x21
   Switch "Interruptor_6" at 267,305 size 40x40

screen "MTA-CompALTA" 1280x800, template "Plantilla"
   GraphicIOField "Plantilla_Campo ES gráfico_3" at 758,425 size 65x60
   GraphicIOField "Plantilla_Campo ES gráfico_4" at 685,353 size 65x60
   GraphicIOField "Plantilla_Campo ES gráfico_5" at 612,281 size 65x60
   GraphicIOField "Plantilla_Campo ES gráfico_2" at 539,209 size 65x60
   GraphicView "Visor de gráficos_2" at 492,46 size 254x172
   GraphicView "Visor de gráficos_18" at 492,46 size 254x172
   GraphicIOField "Plantilla_Campo ES gráfico_1" at 490,113 size 100x102
   GraphicView "Visor de gráficos_3" at 569,134 size 246x148
   ScreenModuleView "Faceplate_8_1" at 781,145 size 47x30
   GraphicView "Visor de gráficos_8" at 1175,577 size 29x50
   GraphicView "Visor de gráficos_7" at 885,605 size 391x113
   TextField "Plantilla_Campo de texto_1" at 1141,578 size 32x23
   IOField "Campo ES_1" at 943,632 size 108x28
   Button "Botón_7" at 1119,186 size 128x41
   Button "Botón_12" at 1119,234 size 128x41
   Button "Botón_13" at 1119,138 size 128x41
   Button "Botón_14" at 641,627 size 160x46
   TextField "Campo de texto_2" at 519,9 size 242x27
   ScreenModuleView "Faceplate_8_5" at 927,289 size 47x30
   ScreenModuleView "Faceplate_8_4" at 1000,361 size 47x30
   GraphicView "Visor de gráficos_19" at 569,134 size 246x148
   ScreenModuleView "Faceplate_8_2" at 854,217 size 47x30
   GraphicView "Visor de gráficos_4" at 642,206 size 246x148
   GraphicView "Visor de gráficos_22" at 642,206 size 246x148
   GraphicView "Visor de gráficos_5" at 715,278 size 246x148
   GraphicView "Visor de gráficos_21" at 715,278 size 246x148
   GraphicView "Visor de gráficos_6" at 788,350 size 246x148
   GraphicView "Visor de gráficos_20" at 788,350 size 246x148
   ScreenModuleView "Faceplate_8_3" at 1072,433 size 47x30
   ScreenModuleView "Faceplate_8_6" at 748,113 size 47x30
   Button "Botón_3" at 1181,68 size 48x46
   ScreenModuleView "Faceplate_8_7" at 1144,505 size 47x30
   GraphicIOField "Plantilla_Campo ES gráfico_6" at 831,497 size 65x60
   GraphicView "Visor de gráficos_1" at 861,422 size 246x148
   GraphicView "Visor de gráficos_9" at 861,422 size 246x148
   GraphicIOField "Campo ES gráfico_4" at 6,182 size 374x6
   SymbolicIOField "Campo ES simbólico_4" at 25,154 size 178x21
   TextField "Campo de texto_1" at 19,121 size 55x32
   GraphicIOField "Campo ES gráfico_5" at 118,341 size 374x6
   TextField "Campo de texto_6" at 127,280 size 67x32
   SymbolicIOField "Campo ES simbólico_5" at 137,313 size 186x21
   GraphicIOField "Campo ES gráfico_1" at 191,422 size 374x6
   TextField "Campo de texto_8" at 200,361 size 67x32
   SymbolicIOField "Campo ES simbólico_1" at 210,394 size 186x21
   GraphicIOField "Campo ES gráfico_3" at 44,262 size 373x6
   TextField "Campo de texto_10" at 53,201 size 67x32
   SymbolicIOField "Campo ES simbólico_3" at 63,234 size 194x21
   GraphicIOField "Campo ES gráfico_2" at 264,502 size 374x6
   TextField "Campo de texto_9" at 273,441 size 67x32
   SymbolicIOField "Campo ES simbólico_2" at 283,474 size 186x21
   GraphicIOField "Campo ES gráfico_16" at 337,582 size 374x6
   TextField "Campo de texto_3" at 346,521 size 67x32
   SymbolicIOField "Campo ES simbólico_11" at 356,554 size 186x21
   IOField "Campo ES_6" at 255,157 size 85x19
   IOField "Campo ES_2" at 367,316 size 85x19
   IOField "Campo ES_3" at 439,397 size 85x19
   IOField "Campo ES_5" at 292,237 size 85x19
   IOField "Campo ES_4" at 512,477 size 85x19
   IOField "Campo ES_7" at 585,557 size 85x19
   ScreenModuleView "Faceplate_6_1" at 283,125 size 57x28
   ScreenModuleView "Faceplate_6_5" at 395,284 size 57x28
   ScreenModuleView "Faceplate_6_4" at 468,365 size 57x28
   ScreenModuleView "Faceplate_6_2" at 321,205 size 57x28
   ScreenModuleView "Faceplate_6_3" at 541,445 size 57x28
   GraphicIOField "Campo ES gráfico_6" at 348,125 size 9x45
   GraphicIOField "Campo ES gráfico_9" at 357,125 size 9x45
   SymbolicIOField "Campo ES simbólico_6" at 86,124 size 160x29
   Button "Botón_11" at 6,116 size 374x64
   Switch "Interruptor_1" at 250,125 size 29x29
   Switch "Interruptor_10" at 863,114 size 40x40
   GraphicIOField "Campo ES gráfico_14" at 459,286 size 9x45
   GraphicIOField "Campo ES gráfico_15" at 468,286 size 9x45
   SymbolicIOField "Campo ES simbólico_10" at 195,283 size 160x29
   Button "Botón_6" at 118,275 size 374x64
   Switch "Interruptor_5" at 360,285 size 29x29
   Switch "Interruptor_9" at 1009,258 size 40x40
   GraphicIOField "Campo ES gráfico_12" at 532,367 size 9x45
   GraphicIOField "Campo ES gráfico_13" at 541,367 size 9x45
   SymbolicIOField "Campo ES simbólico_9" at 269,364 size 160x29
   Button "Botón_8" at 191,356 size 374x64
   Switch "Interruptor_4" at 433,366 size 29x29
   Switch "Interruptor_8" at 1082,330 size 40x40
   GraphicIOField "Campo ES gráfico_7" at 385,207 size 9x45
   GraphicIOField "Campo ES gráfico_10" at 394,207 size 9x45
   SymbolicIOField "Campo ES simbólico_7" at 120,204 size 160x29
   Switch "Interruptor_6" at 936,186 size 40x40
   GraphicIOField "Campo ES gráfico_8" at 605,447 size 9x45
   GraphicIOField "Campo ES gráfico_11" at 614,447 size 9x45
   SymbolicIOField "Campo ES simbólico_8" at 341,444 size 160x29
   Button "Botón_9" at 264,436 size 374x64
   Switch "Interruptor_3" at 504,445 size 29x29
   Switch "Interruptor_7" at 1155,402 size 40x40
   Switch "Interruptor_11" at 1228,474 size 40x40
   ScreenModuleView "Faceplate_6_6" at 614,525 size 57x28
   GraphicIOField "Campo ES gráfico_17" at 678,527 size 9x45
   GraphicIOField "Campo ES gráfico_18" at 687,527 size 9x45
   SymbolicIOField "Campo ES simbólico_12" at 414,524 size 160x29
   Button "Botón_1" at 337,516 size 374x64
   Switch "Interruptor_12" at 577,525 size 29x29
   Button "Botón_10" at 45,196 size 374x64
   Switch "Interruptor_2" at 284,206 size 29x29
   TextField "Campo de texto_4" at 27,564 size 212x67
   IOField "Campo ES_8" at 83,495 size 96x32

